screen "Dos" 800x480, template "Main"
   Button "Button_1" at 7,5 size 96x32; TextOff 'Мешалки'; Authorization "Admin"
      on Release: ActivateScreen("Mix", 0); SetTag("settings", 1)
      Appearance <- "settings"
   Button "Button_2" at 7,52 size 96x32; TextOff 'Дозаторы'; Authorization "Admin"
      on Release: ActivateScreen("Dos", 0); SetTag("settings", 2)
      Appearance <- "settings"
   Button "Button_3" at 7,99 size 96x32; TextOff 'Клапана'; Authorization "Admin"
      on Release: ActivateScreen("Valve", 0); SetTag("settings", 3)
      Appearance <- "settings"
   Button "Button_4" at 7,146 size 96x32; TextOff 'AI'; Authorization "Admin"
      on Release: ActivateScreen("AI", 0); SetTag("settings", 4)
      Appearance <- "settings"
   Button "Button_5" at 7,193 size 96x32; TextOff 'DI'; Authorization "Admin"
      on Release: ActivateScreen("DI", 0); SetTag("settings", 5)
      Appearance <- "settings"
   Button "Button_6" at 7,240 size 96x32; TextOff 'DO'; Authorization "Admin"
      on Release: ActivateScreen("DO", 0); SetTag("settings", 6)
      Appearance <- "settings"
   Group "Group" at 127,7 size 416x126; TextList "Hand"; Picture "z2use_3"; PictureList "Motor"; Text 'Мешалка 1'
   Group "Group_1" at 127,146 size 416x126; Text 'Мешалка 1'; PictureList "Motor"; TextList "Hand"; Picture "z2use_3"
   Group "Group_2" at 127,285 size 416x126; Text 'Мешалка 1'; PictureList "Motor"; TextList "Hand"; Picture "z2use_3"
   Rectangle "Rectangle_1" at 127,7 size 416x126
      Appearance <- "Motors_DB_DD_CMD_Sim"
   GraphicIOField "Graphic I/O field_2" at 134,43 size 43x85; PictureList "Motor"
      ProcessValue <- "Motors_DB_DD_Status"
   Button "Button_7" at 213,41 size 90x22; TextOff 'Авто'; TextList "Hand"
      on Click: InvertBit("Motors_DB_DD_CMD_Hand")
      Appearance <- "Motors_DB_DD_CMD_Hand"
      ProcessValue <- "Motors_DB_DD_CMD_Hand"
   Button "Button_8" at 258,63 size 45x22; TextOff 'Выкл'
      on Click: ResetBit("Motors_DB_DD_CMD_Start_M")
   Button "Button_9" at 213,86 size 90x20; TextOff 'Сервис'
      on Click: InvertBit("Motors_DB_DD_CMD_Service")
      Appearance <- "Motors_DB_DD_CMD_Service"
   Button "Button_13" at 213,63 size 45x22; TextOff 'Вкл'
      on Click: SetBit("Motors_DB_DD_CMD_Start_M")
      Appearance <- "Motors_DB_DD_CMD_Start_M"
   TextField "Text field_13" at 133,12 size 171x26; Text 'Сухой дозатор'
   TextField "Text field_15" at 310,12 size 99x18; Text 'Ожидание ОС, с'
   GraphicView "Graphic view_1" at 180,42 size 25x25; Picture "z2use_3"
      Visibility <- "Motors_DB_DD_CMD_Hand"
   GraphicView "Graphic view_8" at 180,74 size 25x25; Picture "force"
      Visibility <- "Motors_DB_DD_CMD_Force"
   GraphicView "Graphic view_11" at 180,103 size 25x25; Picture "service"
      Visibility <- "Motors_DB_DD_CMD_Service"
   TextField "Text field_3" at 436,31 size 20x18; Text 'QF'
   TextField "Text field_10" at 436,56 size 21x18; Text 'KM'
   TextField "Text field_12" at 436,82 size 44x18; Text 'Service'
   TextField "Text field_14" at 436,108 size 41x18; Text 'Termo'
   TextField "Text field_4" at 416,10 size 120x22; Text 'Использовать:'
   Button "Button_21" at 478,32 size 60x20; TextOff 'Text'; Authorization "Operator"; PictureList "ON_OFF"
      on Click: InvertBit("Motors_DB_DD_Use_QF")
      ProcessValue <- "Motors_DB_DD_Use_QF"
   Button "Button_22" at 478,56 size 60x20; TextOff 'Text'; PictureList "ON_OFF"; Authorization "Operator"
      on Click: InvertBit("Motors_DB_DD_Use_KM")
      ProcessValue <- "Motors_DB_DD_Use_KM"
   Button "Button_24" at 478,80 size 60x20; TextOff 'Text'; PictureList "ON_OFF"; Authorization "Operator"
      on Click: InvertBit("Motors_DB_DD_Use_Serivce")
      ProcessValue <- "Motors_DB_DD_Use_Serivce"
   Button "Button_25" at 478,105 size 60x20; TextOff 'Text'; PictureList "ON_OFF"; Authorization "Operator"
      on Click: InvertBit("Motors_DB_DD_Use_Termo")
      ProcessValue <- "Motors_DB_DD_Use_Termo"
   Button "Button_26" at 416,31 size 20x20; TextOff 'Text'; Authorization "Operator"; PictureList "ok"
      ProcessValue <- "Motors_DB_DD_FB_QF"
   Button "Button_27" at 416,55 size 20x20; TextOff 'Text'; PictureList "ok"; Authorization "Operator"
      ProcessValue <- "Motors_DB_DD_FB_KM"
   Button "Button_29" at 416,80 size 20x20; TextOff 'Text'; PictureList "ok"; Authorization "Operator"
      ProcessValue <- "Motors_DB_DD_Use_Serivce"
   Button "Button_30" at 416,105 size 20x20; TextOff 'Text'; PictureList "ok"; Authorization "Operator"
      ProcessValue <- "Motors_DB_DD_FB_Termo"
   TextField "Text field_1" at 323,87 size 79x18; Text 'Наработка, ч'
   TextField "Text field_2" at 309,34 size 37x18; Text 'Старт'
   IOField "I/O field_5" at 348,32 size 30x20; FormatPattern 99
      ProcessValue <- "Motors_DB_DD_Wait_On_SP"
   IOField "I/O field_12" at 348,55 size 30x20; FormatPattern 99
      ProcessValue <- "Motors_DB_DD_Wait_Off_SP"
   TextField "Text field_5" at 309,55 size 32x18; Text 'Стоп'
   IOField "I/O field_13" at 378,32 size 30x20; FormatPattern 99
      ProcessValue <- "Motors_DB_DD_Wait_On_Now"
   IOField "I/O field_14" at 378,55 size 30x20; FormatPattern 99
      ProcessValue <- "Motors_DB_DD_Wait_Off_Now"
   IOField "I/O field_16" at 313,105 size 98x20; FormatPattern 9999999999
      ProcessValue <- "Motors_DB_DD_Res_h"
   Button "Button_11" at 213,106 size 90x20; TextOff 'Force'
      on Click: InvertBit("Motors_DB_DD_CMD_Force")
      Appearance <- "Motors_DB_DD_CMD_Force"
   Rectangle "Rectangle_2" at 127,146 size 416x126
      Appearance <- "Motors_DB_Vibro_CMD_Sim"
   GraphicIOField "Graphic I/O field_1" at 134,182 size 43x85; PictureList "Motor"
      ProcessValue <- "Motors_DB_Vibro_Status"
   Button "Button_10" at 213,180 size 90x22; TextOff 'Авто'; TextList "Hand"
      on Click: InvertBit("Motors_DB_Vibro_CMD_Hand")
      Appearance <- "Motors_DB_Vibro_CMD_Hand"
      ProcessValue <- "Motors_DB_Vibro_CMD_Hand"
   Button "Button_12" at 258,202 size 45x22; TextOff 'Выкл'
      on Click: ResetBit("Motors_DB_Vibro_CMD_Start_M")
   Button "Button_14" at 213,225 size 90x20; TextOff 'Сервис'
      on Click: InvertBit("Motors_DB_Vibro_CMD_Service")
      Appearance <- "Motors_DB_Vibro_CMD_Service"
   Button "Button_15" at 213,202 size 45x22; TextOff 'Вкл'
      on Click: SetBit("Motors_DB_Vibro_CMD_Start_M")
      Appearance <- "Motors_DB_Vibro_CMD_Start_M"
   TextField "Text field_6" at 133,151 size 171x26; Text 'Вибратор'
   TextField "Text field_7" at 310,151 size 99x18; Text 'Ожидание ОС, с'
   GraphicView "Graphic view_2" at 180,181 size 25x25; Picture "z2use_3"
      Visibility <- "Motors_DB_Vibro_CMD_Hand"
   GraphicView "Graphic view_3" at 180,213 size 25x25; Picture "force"
      Visibility <- "Motors_DB_Vibro_CMD_Force"
   GraphicView "Graphic view_4" at 180,242 size 25x25; Picture "service"
      Visibility <- "Motors_DB_Vibro_CMD_Service"
   TextField "Text field_8" at 436,170 size 20x18; Text 'QF'
   TextField "Text field_9" at 436,195 size 21x18; Text 'KM'
   TextField "Text field_11" at 436,221 size 44x18; Text 'Service'
   TextField "Text field_16" at 436,247 size 41x18; Text 'Termo'
   TextField "Text field_17" at 416,149 size 120x22; Text 'Использовать:'
   Button "Button_16" at 478,171 size 60x20; TextOff 'Text'; PictureList "ON_OFF"; Authorization "Operator"
      on Click: InvertBit("Motors_DB_Vibro_Use_QF")
      ProcessValue <- "Motors_DB_Vibro_Use_QF"
   Button "Button_17" at 478,195 size 60x20; TextOff 'Text'; Authorization "Operator"; PictureList "ON_OFF"
      on Click: InvertBit("Motors_DB_Vibro_Use_KM")
      ProcessValue <- "Motors_DB_Vibro_Use_KM"
   Button "Button_18" at 478,219 size 60x20; TextOff 'Text'; Authorization "Operator"; PictureList "ON_OFF"
      on Click: InvertBit("Motors_DB_Vibro_Use_Serivce")
      ProcessValue <- "Motors_DB_Vibro_Use_Serivce"
   Button "Button_19" at 478,244 size 60x20; TextOff 'Text'; Authorization "Operator"; PictureList "ON_OFF"
      on Click: InvertBit("Motors_DB_Vibro_Use_Termo")
      ProcessValue <- "Motors_DB_Vibro_Use_Termo"
   Button "Button_20" at 416,170 size 20x20; TextOff 'Text'; PictureList "ok"; Authorization "Operator"
      ProcessValue <- "Motors_DB_Vibro_FB_QF"
   Button "Button_23" at 416,194 size 20x20; TextOff 'Text'; Authorization "Operator"; PictureList "ok"
      ProcessValue <- "Motors_DB_Vibro_FB_KM"
   Button "Button_28" at 416,219 size 20x20; TextOff 'Text'; Authorization "Operator"; PictureList "ok"
      ProcessValue <- "Motors_DB_Vibro_Use_Serivce"
   Button "Button_31" at 416,244 size 20x20; TextOff 'Text'; Authorization "Operator"; PictureList "ok"
      ProcessValue <- "Motors_DB_Vibro_FB_Termo"
   TextField "Text field_18" at 323,226 size 79x18; Text 'Наработка, ч'
   TextField "Text field_19" at 309,173 size 37x18; Text 'Старт'
   IOField "I/O field_1" at 348,171 size 30x20; FormatPattern 99
      ProcessValue <- "Motors_DB_Vibro_Wait_On_SP"
   IOField "I/O field_2" at 348,194 size 30x20; FormatPattern 99
      ProcessValue <- "Motors_DB_Vibro_Wait_Off_SP"
   TextField "Text field_20" at 309,194 size 32x18; Text 'Стоп'
   IOField "I/O field_3" at 378,171 size 30x20; FormatPattern 99
      ProcessValue <- "Motors_DB_Vibro_Wait_On_Now"
   IOField "I/O field_4" at 378,194 size 30x20; FormatPattern 99
      ProcessValue <- "Motors_DB_Vibro_Wait_Off_Now"
   IOField "I/O field_6" at 313,244 size 98x20; FormatPattern 9999999999
      ProcessValue <- "Motors_DB_Vibro_Res_h"
   Button "Button_32" at 213,245 size 90x20; TextOff 'Force'
      on Click: InvertBit("Motors_DB_Vibro_CMD_Force")
      Appearance <- "Motors_DB_Vibro_CMD_Force"
   Rectangle "Rectangle_3" at 127,285 size 416x126
      Appearance <- "Motors_DB_DL_CMD_Sim"
   GraphicIOField "Graphic I/O field_3" at 134,321 size 43x85; PictureList "Motor"
      ProcessValue <- "Motors_DB_DL_Status"
   Button "Button_33" at 213,319 size 90x22; TextOff 'Авто'; TextList "Hand"
      on Click: InvertBit("Motors_DB_DL_CMD_Hand")
      Appearance <- "Motors_DB_DL_CMD_Hand"
      ProcessValue <- "Motors_DB_DL_CMD_Hand"
   Button "Button_34" at 258,341 size 45x22; TextOff 'Выкл'
      on Click: ResetBit("Motors_DB_DL_CMD_Start_M")
   Button "Button_35" at 213,364 size 90x20; TextOff 'Сервис'
      on Click: InvertBit("Motors_DB_DL_CMD_Service")
      Appearance <- "Motors_DB_DL_CMD_Service"
   Button "Button_36" at 213,341 size 45x22; TextOff 'Вкл'
      on Click: SetBit("Motors_DB_DL_CMD_Start_M")
      Appearance <- "Motors_DB_DL_CMD_Start_M"
   TextField "Text field_21" at 133,290 size 171x26; Text 'Жидкий дозатор'
   TextField "Text field_22" at 310,290 size 99x18; Text 'Ожидание ОС, с'
   GraphicView "Graphic view_5" at 180,320 size 25x25; Picture "z2use_3"
      Visibility <- "Motors_DB_DL_CMD_Hand"
   GraphicView "Graphic view_6" at 180,352 size 25x25; Picture "force"
      Visibility <- "Motors_DB_DL_CMD_Force"
   GraphicView "Graphic view_7" at 180,381 size 25x25; Picture "service"
      Visibility <- "Motors_DB_DL_CMD_Service"
   TextField "Text field_23" at 436,309 size 20x18; Text 'QF'
   TextField "Text field_24" at 436,334 size 21x18; Text 'KM'
   TextField "Text field_25" at 436,360 size 44x18; Text 'Service'
   TextField "Text field_26" at 436,386 size 41x18; Text 'Termo'
   TextField "Text field_27" at 416,288 size 120x22; Text 'Использовать:'
   Button "Button_37" at 478,310 size 60x20; TextOff 'Text'; PictureList "ON_OFF"; Authorization "Operator"
      on Click: InvertBit("Motors_DB_DL_Use_QF")
      ProcessValue <- "Motors_DB_DL_Use_QF"
   Button "Button_38" at 478,334 size 60x20; TextOff 'Text'; Authorization "Operator"; PictureList "ON_OFF"
      on Click: InvertBit("Motors_DB_DL_Use_KM")
      ProcessValue <- "Motors_DB_DL_Use_KM"
   Button "Button_39" at 478,358 size 60x20; TextOff 'Text'; Authorization "Operator"; PictureList "ON_OFF"
      on Click: InvertBit("Motors_DB_DL_Use_Serivce")
      ProcessValue <- "Motors_DB_DL_Use_Serivce"
   Button "Button_40" at 478,383 size 60x20; TextOff 'Text'; Authorization "Operator"; PictureList "ON_OFF"
      on Click: InvertBit("Motors_DB_DL_Use_Termo")
      ProcessValue <- "Motors_DB_DL_Use_Termo"
   Button "Button_41" at 416,309 size 20x20; TextOff 'Text'; PictureList "ok"; Authorization "Operator"
      ProcessValue <- "Motors_DB_DL_FB_QF"
   Button "Button_42" at 416,333 size 20x20; TextOff 'Text'; Authorization "Operator"; PictureList "ok"
      ProcessValue <- "Motors_DB_DL_FB_KM"
   Button "Button_43" at 416,358 size 20x20; TextOff 'Text'; Authorization "Operator"; PictureList "ok"
      ProcessValue <- "Motors_DB_DL_Use_Serivce"
   Button "Button_44" at 416,383 size 20x20; TextOff 'Text'; Authorization "Operator"; PictureList "ok"
      ProcessValue <- "Motors_DB_DL_FB_Termo"
   TextField "Text field_28" at 323,365 size 79x18; Text 'Наработка, ч'
   TextField "Text field_29" at 309,312 size 37x18; Text 'Старт'
   IOField "I/O field_7" at 348,310 size 30x20; FormatPattern 99
      ProcessValue <- "Motors_DB_DL_Wait_On_SP"
   IOField "I/O field_8" at 348,333 size 30x20; FormatPattern 99
      ProcessValue <- "Motors_DB_DL_Wait_Off_SP"
   TextField "Text field_30" at 309,333 size 32x18; Text 'Стоп'
   IOField "I/O field_9" at 378,310 size 30x20; FormatPattern 99
      ProcessValue <- "Motors_DB_DL_Wait_On_Now"
   IOField "I/O field_10" at 378,333 size 30x20; FormatPattern 99
      ProcessValue <- "Motors_DB_DL_Wait_Off_Now"
   IOField "I/O field_11" at 313,383 size 98x20; FormatPattern 9999999999
      ProcessValue <- "Motors_DB_DL_Res_h"
   Button "Button_45" at 213,384 size 90x20; TextOff 'Force'
      on Click: InvertBit("Motors_DB_DL_CMD_Force")
      Appearance <- "Motors_DB_DL_CMD_Force"

screen "Valve" 800x480, template "Main"
   Button "Button_1" at 7,5 size 96x32; TextOff 'Мешалки'; Authorization "Admin"
      on Release: ActivateScreen("Mix", 0); SetTag("settings", 1)
      Appearance <- "settings"
   Button "Button_2" at 7,52 size 96x32; TextOff 'Дозаторы'; Authorization "Admin"
      on Release: ActivateScreen("Dos", 0); SetTag("settings", 2)
      Appearance <- "settings"
   Button "Button_3" at 7,99 size 96x32; TextOff 'Клапана'; Authorization "Admin"
      on Release: ActivateScreen("Valve", 0); SetTag("settings", 3)
      Appearance <- "settings"
   Button "Button_4" at 7,146 size 96x32; TextOff 'AI'; Authorization "Admin"
      on Release: ActivateScreen("AI", 0); SetTag("settings", 4)
      Appearance <- "settings"
   Button "Button_5" at 7,193 size 96x32; TextOff 'DI'; Authorization "Admin"
      on Release: ActivateScreen("DI", 0); SetTag("settings", 5)
      Appearance <- "settings"
   Button "Button_6" at 7,240 size 96x32; TextOff 'DO'; Authorization "Admin"
      on Release: ActivateScreen("DO", 0); SetTag("settings", 6)
      Appearance <- "settings"
   Group "Group" at 127,7 size 264x51; TextList "Hand"
   Rectangle "Rectangle_2" at 127,7 size 264x51
      Appearance <- "Micro_DB_KC1_Alarm"
   TextField "Text field_5" at 130,10 size 97x22; Text 'Клапан КС1'
   Button "Button_13" at 246,11 size 59x44; TextOff 'Авто'; TextList "Hand"
      on Click: InvertBit("Micro_DB_KC1_Hand")
      Appearance <- "Micro_DB_KC1_Hand"
      ProcessValue <- "Micro_DB_KC1_Hand"
   Button "Button_14" at 188,33 size 49x22; TextOff 'Выкл'
      on Click: ResetBit("Micro_DB_KC1_Start_M")
   Button "Button_15" at 132,33 size 47x22; TextOff 'Вкл'
      on Click: SetBit("Micro_DB_KC1_Start_M")
      Appearance <- "Micro_DB_KC1_Start_M"
   TextField "Text field_1" at 306,8 size 28x23; Text 'ОС'
   Button "Button_7" at 336,11 size 50x20; TextOff 'Text'; Authorization "Operator"; PictureList "ON_OFF"
      on Click: InvertBit("Micro_DB_KC1_No_FB")
      ProcessValue <- "Micro_DB_KC1_No_FB"
   IOField "I/O field_5" at 308,31 size 30x22; FormatPattern 99
      ProcessValue <- "Micro_DB_KC1_Wait_On_SP"
   IOField "I/O field_8" at 355,31 size 30x22; FormatPattern 99
      ProcessValue <- "Micro_DB_KC1_Wait_Off_SP"

screen "AI" 800x480, template "Main"
   Button "Button_1" at 7,5 size 96x32; TextOff 'Мешалки'; Authorization "Admin"
      on Release: ActivateScreen("Mix", 0); SetTag("settings", 1)
      Appearance <- "settings"
   Button "Button_2" at 7,52 size 96x32; TextOff 'Дозаторы'; Authorization "Admin"
      on Release: ActivateScreen("Dos", 0); SetTag("settings", 2)
      Appearance <- "settings"
   Button "Button_3" at 7,99 size 96x32; TextOff 'Клапана'; Authorization "Admin"
      on Release: ActivateScreen("Valve", 0); SetTag("settings", 3)
      Appearance <- "settings"
   Button "Button_4" at 7,146 size 96x32; TextOff 'AI'; Authorization "Admin"
      on Release: ActivateScreen("AI", 0); SetTag("settings", 4)
      Appearance <- "settings"
   Button "Button_5" at 7,193 size 96x32; TextOff 'DI'; Authorization "Admin"
      on Release: ActivateScreen("DI", 0); SetTag("settings", 5)
      Appearance <- "settings"
   Button "Button_6" at 7,240 size 96x32; TextOff 'DO'; Authorization "Admin"
      on Release: ActivateScreen("DO", 0); SetTag("settings", 6)
      Appearance <- "settings"
   TextField "Text field_2" at 210,15 size 67x22; Text 'Датчик:'
   TextField "Text field_4" at 282,15 size 99x22; Text 'Расходомер'
   TextField "Text field_7" at 390,18 size 43x22; Text 'вход'
   TextField "Text field_8" at 390,43 size 56x22; Text 'выход'
   IOField "I/O field_1" at 456,19 size 92x26; FormatPattern s999999999.999
      ProcessValue <- "AIx_DB_FlowMeter_Converter_Min_In"
   IOField "I/O field_2" at 456,41 size 92x26; FormatPattern s999999999.999
      ProcessValue <- "AIx_DB_FlowMeter_Converter_Min_Out"
   IOField "I/O field_3" at 555,18 size 92x26; FormatPattern s999999999.999
      ProcessValue <- "AIx_DB_FlowMeter_Converter_Max_In"
   IOField "I/O field_4" at 555,40 size 92x26; FormatPattern s999999999.999
      ProcessValue <- "AIx_DB_FlowMeter_Converter_Max_Out"
   TextField "Text field_9" at 389,68 size 101x22; Text 'Фильтрация'
   TextField "Text field_10" at 390,96 size 36x22; Text 'RTD'
   Button "Button_7" at 489,71 size 20x20; TextOff 'Text'; PictureList "ok"
      ProcessValue <- "AIx_DB_FlowMeter_Use_Filter"
      on Click: InvertBit("AIx_DB_FlowMeter_Use_Filter")
   Button "Button_8" at 489,96 size 20x20; TextOff 'Text'; PictureList "ok"
      on Click: InvertBit("AIx_DB_FlowMeter_Use_RTD")
      ProcessValue <- "AIx_DB_FlowMeter_Use_RTD"
   IOField "I/O field_5" at 516,68 size 65x25; FormatPattern 999
      ProcessValue <- "AIx_DB_FlowMeter_Filter_SP"
   IOField "I/O field_6" at 516,93 size 65x25; FormatPattern 999
      ProcessValue <- "AIx_DB_FlowMeter_RTD_c"
   TextField "Text field_11" at 210,36 size 79x22; Text 'Поправка'
   IOField "I/O field_7" at 293,36 size 78x23; FormatPattern s999.9
      ProcessValue <- "AIx_DB_FlowMeter_Calibration"
   Button "Button_9" at 396,176 size 248x28; TextOff 'Use'
      Appearance <- "AIx_DB_FlowMeter_CMD_Start_A"
      on Click: InvertBit("AIx_DB_FlowMeter_CMD_Start_A")
   Button "Button_10" at 213,66 size 68x28; TextOff 'Hand'
      on Click: InvertBit("AIx_DB_FlowMeter_CMD_Hand")
      Appearance <- "AIx_DB_FlowMeter_CMD_Hand"
   IOField "I/O field_8" at 293,66 size 78x28; FormatPattern s9999.9
      ProcessValue <- "AIx_DB_FlowMeter_Result"
   TextField "Text field_12" at 436,123 size 27x22; Text 'NC'
   TextField "Text field_13" at 437,143 size 25x22; Text 'SC'
   TextField "Text field_14" at 210,125 size 27x22; Text 'HH'
   TextField "Text field_15" at 216,145 size 16x22; Text 'H'
   TextField "Text field_16" at 217,165 size 14x22; Text 'L'
   TextField "Text field_17" at 212,186 size 23x22; Text 'LL'
   IOField "I/O field_11" at 472,123 size 58x21; FormatPattern s99999
      ProcessValue <- "AIx_DB_FlowMeter_SP_NC"
   IOField "I/O field_12" at 472,143 size 58x21; FormatPattern s99999
      ProcessValue <- "AIx_DB_FlowMeter_SP_SC"
   IOField "I/O field_13" at 246,125 size 58x21; FormatPattern 99999
      ProcessValue <- "AIx_DB_FlowMeter_SP_HH"
   IOField "I/O field_14" at 246,145 size 58x21; FormatPattern 99999
      ProcessValue <- "AIx_DB_FlowMeter_SP_H"
   IOField "I/O field_15" at 246,165 size 58x21; FormatPattern s99999
      ProcessValue <- "AIx_DB_FlowMeter_SP_L"
   IOField "I/O field_16" at 246,185 size 58x21; FormatPattern s99999
      ProcessValue <- "AIx_DB_FlowMeter_SP_LL"
   IOField "I/O field_17" at 546,123 size 58x21; FormatPattern 999
      ProcessValue <- "AIx_DB_FlowMeter_Timers_NC_SP"
   IOField "I/O field_18" at 546,143 size 58x21; FormatPattern 999
      ProcessValue <- "AIx_DB_FlowMeter_Timers_SC_SP"
   IOField "I/O field_19" at 320,125 size 58x21; FormatPattern 999
      ProcessValue <- "AIx_DB_FlowMeter_Timers_HH_SP"
   IOField "I/O field_20" at 320,145 size 58x21; FormatPattern 999
      ProcessValue <- "AIx_DB_FlowMeter_Timers_H_SP"
   IOField "I/O field_21" at 320,165 size 58x21; FormatPattern 999
      ProcessValue <- "AIx_DB_FlowMeter_Timers_L_SP"
   IOField "I/O field_22" at 320,185 size 58x21; FormatPattern 999
      ProcessValue <- "AIx_DB_FlowMeter_Timers_LL_SP"
   IOField "I/O field_23" at 582,93 size 65x25; FormatPattern s99999
      ProcessValue <- "AIx_DB_FlowMeter_Signal"
   TextField "Text field_18" at 210,97 size 68x22; Text 'Уставка'
   TextField "Text field_19" at 299,97 size 79x22; Text 'Время (с)'
   TextField "Text field_1" at 214,248 size 67x22; Text 'Датчик:'
   TextField "Text field_3" at 286,248 size 69x22; Text 'Уровень'
   TextField "Text field_5" at 394,251 size 43x22; Text 'вход'
   TextField "Text field_6" at 394,276 size 56x22; Text 'выход'
   IOField "I/O field_9" at 460,252 size 92x26; FormatPattern s999999999.999
      ProcessValue <- "AIx_DB_Level_Converter_Min_In"
   IOField "I/O field_10" at 460,274 size 92x26; FormatPattern s999999999.999
      ProcessValue <- "AIx_DB_Level_Converter_Min_Out"
   IOField "I/O field_24" at 559,251 size 92x26; FormatPattern s999999999.999
      ProcessValue <- "AIx_DB_Level_Converter_Max_In"
   IOField "I/O field_25" at 559,273 size 92x26; FormatPattern s999999999.999
      ProcessValue <- "AIx_DB_Level_Converter_Max_Out"
   TextField "Text field_20" at 393,301 size 101x22; Text 'Фильтрация'
   TextField "Text field_21" at 394,329 size 36x22; Text 'RTD'
   Button "Button_11" at 493,304 size 20x20; TextOff 'Text'; PictureList "ok"
      on Click: InvertBit("AIx_DB_Level_Use_Filter")
      ProcessValue <- "AIx_DB_Level_Use_Filter"
   Button "Button_12" at 493,329 size 20x20; TextOff 'Text'; PictureList "ok"
      on Click: InvertBit("AIx_DB_Level_Use_RTD")
      ProcessValue <- "AIx_DB_Level_Use_RTD"
   IOField "I/O field_26" at 520,301 size 65x25; FormatPattern 999
      ProcessValue <- "AIx_DB_Level_Filter_SP"
   IOField "I/O field_27" at 520,326 size 65x25; FormatPattern 999
      ProcessValue <- "AIx_DB_Level_RTD_c"
   TextField "Text field_22" at 214,269 size 79x22; Text 'Поправка'
   IOField "I/O field_28" at 297,269 size 78x23; FormatPattern s999.9
      ProcessValue <- "AIx_DB_Level_Calibration"
   Button "Button_13" at 400,409 size 248x28; TextOff 'Use'
      on Click: InvertBit("AIx_DB_Level_CMD_Start_A")
      Appearance <- "AIx_DB_Level_CMD_Start_A"
   Button "Button_14" at 217,299 size 68x28; TextOff 'Hand'
      on Click: InvertBit("AIx_DB_Level_CMD_Hand")
      Appearance <- "AIx_DB_Level_CMD_Hand"
   IOField "I/O field_29" at 297,299 size 78x28; FormatPattern s9999.9
      ProcessValue <- "AIx_DB_Level_Result"
   TextField "Text field_23" at 440,356 size 27x22; Text 'NC'
   TextField "Text field_24" at 441,376 size 25x22; Text 'SC'
   TextField "Text field_25" at 214,358 size 27x22; Text 'HH'
   TextField "Text field_26" at 220,378 size 16x22; Text 'H'
   TextField "Text field_27" at 221,398 size 14x22; Text 'L'
   TextField "Text field_28" at 216,419 size 23x22; Text 'LL'
   IOField "I/O field_30" at 476,356 size 58x21; FormatPattern s99999
      ProcessValue <- "AIx_DB_Level_SP_NC"
   IOField "I/O field_31" at 476,376 size 58x21; FormatPattern s99999
      ProcessValue <- "AIx_DB_Level_SP_SC"
   IOField "I/O field_32" at 250,358 size 58x21; FormatPattern 99999
      ProcessValue <- "AIx_DB_Level_SP_HH"
   IOField "I/O field_33" at 250,378 size 58x21; FormatPattern 99999
      ProcessValue <- "AIx_DB_Level_SP_H"
   IOField "I/O field_34" at 250,398 size 58x21; FormatPattern s99999
      ProcessValue <- "AIx_DB_Level_SP_L"
   IOField "I/O field_35" at 250,418 size 58x21; FormatPattern s99999
      ProcessValue <- "AIx_DB_Level_SP_LL"
   IOField "I/O field_36" at 550,356 size 58x21; FormatPattern 999
      ProcessValue <- "AIx_DB_Level_Timers_NC_SP"
   IOField "I/O field_37" at 550,376 size 58x21; FormatPattern 999
      ProcessValue <- "AIx_DB_Level_Timers_SC_SP"
   IOField "I/O field_38" at 324,358 size 58x21; FormatPattern 999
      ProcessValue <- "AIx_DB_Level_Timers_HH_SP"
   IOField "I/O field_39" at 324,378 size 58x21; FormatPattern 999
      ProcessValue <- "AIx_DB_Level_Timers_H_SP"
   IOField "I/O field_40" at 324,398 size 58x21; FormatPattern 999
      ProcessValue <- "AIx_DB_Level_Timers_L_SP"
   IOField "I/O field_41" at 324,418 size 58x21; FormatPattern 999
      ProcessValue <- "AIx_DB_Level_Timers_LL_SP"
   IOField "I/O field_42" at 586,326 size 65x25; FormatPattern s99999
      ProcessValue <- "AIx_DB_Level_Signal"
   TextField "Text field_29" at 214,330 size 68x22; Text 'Уставка'
   TextField "Text field_30" at 303,330 size 79x22; Text 'Время (с)'

screen "DI" 800x480, template "Main"
   Button "Button_1" at 7,5 size 96x32; TextOff 'Мешалки'; Authorization "Admin"
      on Release: ActivateScreen("Mix", 0); SetTag("settings", 1)
      Appearance <- "settings"
   Button "Button_2" at 7,52 size 96x32; TextOff 'Дозаторы'; Authorization "Admin"
      on Release: ActivateScreen("Dos", 0); SetTag("settings", 2)
      Appearance <- "settings"
   Button "Button_3" at 7,99 size 96x32; TextOff 'Клапана'; Authorization "Admin"
      on Release: ActivateScreen("Valve", 0); SetTag("settings", 3)
      Appearance <- "settings"
   Button "Button_4" at 7,146 size 96x32; TextOff 'AI'; Authorization "Admin"
      on Release: ActivateScreen("AI", 0); SetTag("settings", 4)
      Appearance <- "settings"
   Button "Button_5" at 7,193 size 96x32; TextOff 'DI'; Authorization "Admin"
      on Release: ActivateScreen("DI", 0); SetTag("settings", 5)
      Appearance <- "settings"
   Button "Button_6" at 7,240 size 96x32; TextOff 'DO'; Authorization "Admin"
      on Release: ActivateScreen("DO", 0); SetTag("settings", 6)
      Appearance <- "settings"
   Group "Group" at 127,7 size 283x51; TextList "Hand"
   Group "Group_1" at 127,66 size 283x51; TextList "Hand"
   Group "Group_2" at 127,125 size 283x51; TextList "Hand"
   Group "Group_3" at 127,184 size 283x51; TextList "Hand"
   Group "Group_4" at 127,244 size 283x51; TextList "Hand"
   Group "Group_5" at 127,303 size 283x51; TextList "Hand"
   Group "Group_6" at 127,362 size 283x51; TextList "Hand"
   Group "Group_7" at 127,422 size 283x51; TextList "Hand"
   Group "Group_8" at 433,7 size 283x51; TextList "Hand"
   Group "Group_9" at 433,66 size 283x51; TextList "Hand"
   Group "Group_10" at 433,125 size 283x51; TextList "Hand"
   Group "Group_11" at 433,184 size 283x51; TextList "Hand"
   Group "Group_12" at 433,244 size 283x51; TextList "Hand"
   Group "Group_13" at 433,303 size 283x51; TextList "Hand"
   TextField "Text field_1" at 131,10 size 45x22; Text 'I 0.0'
   TextField "Text field_2" at 176,10 size 120x22; Text 'M1 Готовность'
   Circle "Circle_1" at 131,33 size 22x22
      Appearance <- "DIx_DB_M1_FB_Ready_Input"
   Circle "Circle_2" at 154,33 size 22x22
      Appearance <- "DIx_DB_M1_FB_Ready_Signal"
   Button "Button_7" at 298,11 size 59x44; TextOff 'Авто'; TextList "Hand"
      on Click: InvertBit("DIx_DB_M1_FB_Ready_Hand")
      Appearance <- "DIx_DB_M1_FB_Ready_Hand"
      ProcessValue <- "DIx_DB_M1_FB_Ready_Hand"
   Button "Button_8" at 240,33 size 49x22; TextOff 'Выкл'
      on Click: ResetBit("DIx_DB_M1_FB_Ready_Start_M")
   Button "Button_12" at 184,33 size 47x22; TextOff 'Вкл'
      Appearance <- "DIx_DB_M1_FB_Ready_Start_M"
      on Click: SetBit("DIx_DB_M1_FB_Ready_Start_M")
   IOField "I/O field_6" at 360,33 size 23x22; FormatPattern 99
      ProcessValue <- "DIx_DB_M1_FB_Ready_Filter_On_SP"
   IOField "I/O field_7" at 383,33 size 23x22; FormatPattern 99
      ProcessValue <- "DIx_DB_M1_FB_Ready_Filter_Off_SP"
   Button "Button_9" at 360,10 size 46x20; TextOff 'Inv'
      Appearance <- "DIx_DB_M1_FB_Ready_Inverse"
      on Click: InvertBit("DIx_DB_M1_FB_Ready_Inverse")
   TextField "Text field_3" at 131,69 size 45x22; Text 'I 0.1'
   TextField "Text field_4" at 176,69 size 87x22; Text 'M1 Работа'
   Circle "Circle_3" at 131,92 size 22x22
      Appearance <- "DIx_DB_M1_FB_Run_Input"
   Circle "Circle_4" at 154,92 size 22x22
      Appearance <- "DIx_DB_M1_FB_Run_Signal"
   Button "Button_10" at 298,70 size 59x44; TextOff 'Авто'; TextList "Hand"
      on Click: InvertBit("DIx_DB_M1_FB_Run_Hand")
      Appearance <- "DIx_DB_M1_FB_Run_Hand"
      ProcessValue <- "DIx_DB_M1_FB_Run_Hand"
   Button "Button_11" at 240,92 size 49x22; TextOff 'Выкл'
      on Click: ResetBit("DIx_DB_M1_FB_Run_Start_M")
   Button "Button_13" at 184,92 size 47x22; TextOff 'Вкл'
      on Click: SetBit("DIx_DB_M1_FB_Run_Start_M")
      Appearance <- "DIx_DB_M1_FB_Run_Start_M"
   IOField "I/O field_1" at 360,92 size 23x22; FormatPattern 99
      ProcessValue <- "DIx_DB_M1_FB_Run_Filter_On_SP"
   IOField "I/O field_2" at 383,92 size 23x22; FormatPattern 99
      ProcessValue <- "DIx_DB_M1_FB_Run_Filter_Off_SP"
   Button "Button_14" at 360,69 size 46x20; TextOff 'Inv'
      on Click: InvertBit("DIx_DB_M1_FB_Run_Inverse")
      Appearance <- "DIx_DB_M1_FB_Run_Inverse"
   TextField "Text field_5" at 131,128 size 45x22; Text 'I 0.2'
   TextField "Text field_6" at 176,128 size 120x22; Text 'M2 Готовность'
   Circle "Circle_5" at 131,151 size 22x22
      Appearance <- "DIx_DB_M2_FB_Ready_Input"
   Circle "Circle_6" at 154,151 size 22x22
      Appearance <- "DIx_DB_M2_FB_Ready_Signal"
   Button "Button_15" at 298,129 size 59x44; TextOff 'Авто'; TextList "Hand"
      on Click: InvertBit("DIx_DB_M2_FB_Ready_Hand")
      Appearance <- "DIx_DB_M2_FB_Ready_Hand"
      ProcessValue <- "DIx_DB_M2_FB_Ready_Hand"
   Button "Button_16" at 240,151 size 49x22; TextOff 'Выкл'
      on Click: ResetBit("DIx_DB_M2_FB_Ready_Start_M")
   Button "Button_17" at 184,151 size 47x22; TextOff 'Вкл'
      on Click: SetBit("DIx_DB_M2_FB_Ready_Start_M")
      Appearance <- "DIx_DB_M2_FB_Ready_Start_M"
   IOField "I/O field_3" at 360,151 size 23x22; FormatPattern 99
      ProcessValue <- "DIx_DB_M2_FB_Ready_Filter_On_SP"
   IOField "I/O field_4" at 383,151 size 23x22; FormatPattern 99
      ProcessValue <- "DIx_DB_M2_FB_Ready_Filter_Off_SP"
   Button "Button_18" at 360,128 size 46x20; TextOff 'Inv'
      on Click: InvertBit("DIx_DB_M2_FB_Ready_Inverse")
      Appearance <- "DIx_DB_M2_FB_Ready_Inverse"
   TextField "Text field_7" at 131,187 size 45x22; Text 'I 0.3'
   TextField "Text field_8" at 176,187 size 87x22; Text 'M2 Работа'
   Circle "Circle_7" at 131,210 size 22x22
      Appearance <- "DIx_DB_M2_FB_Run_Input"
   Circle "Circle_8" at 154,210 size 22x22
      Appearance <- "DIx_DB_M2_FB_Run_Signal"
   Button "Button_19" at 298,188 size 59x44; TextOff 'Авто'; TextList "Hand"
      on Click: InvertBit("DIx_DB_M2_FB_Run_Hand")
      Appearance <- "DIx_DB_M2_FB_Run_Hand"
      ProcessValue <- "DIx_DB_M2_FB_Run_Hand"
   Button "Button_20" at 240,210 size 49x22; TextOff 'Выкл'
      on Click: ResetBit("DIx_DB_M2_FB_Run_Start_M")
   Button "Button_21" at 184,210 size 47x22; TextOff 'Вкл'
      on Click: SetBit("DIx_DB_M2_FB_Run_Start_M")
      Appearance <- "DIx_DB_M2_FB_Run_Start_M"
   IOField "I/O field_5" at 360,210 size 23x22; FormatPattern 99
      ProcessValue <- "DIx_DB_M2_FB_Run_Filter_On_SP"
   IOField "I/O field_8" at 383,210 size 23x22; FormatPattern 99
      ProcessValue <- "DIx_DB_M2_FB_Run_Filter_Off_SP"
   Button "Button_22" at 360,187 size 46x20; TextOff 'Inv'
      on Click: InvertBit("DIx_DB_M2_FB_Run_Inverse")
      Appearance <- "DIx_DB_M2_FB_Run_Inverse"
   TextField "Text field_9" at 131,247 size 45x22; Text 'I 0.4'
   TextField "Text field_10" at 176,247 size 120x22; Text 'M3 Готовность'
   Circle "Circle_9" at 131,270 size 22x22
      Appearance <- "DIx_DB_M3_FB_Ready_Input"
   Circle "Circle_10" at 154,270 size 22x22
      Appearance <- "DIx_DB_M3_FB_Ready_Signal"
   Button "Button_23" at 298,248 size 59x44; TextOff 'Авто'; TextList "Hand"
      on Click: InvertBit("DIx_DB_M3_FB_Ready_Hand")
      Appearance <- "DIx_DB_M3_FB_Ready_Hand"
      ProcessValue <- "DIx_DB_M3_FB_Ready_Hand"
   Button "Button_24" at 240,270 size 49x22; TextOff 'Выкл'
      on Click: ResetBit("DIx_DB_M3_FB_Ready_Start_M")
   Button "Button_25" at 184,270 size 47x22; TextOff 'Вкл'
      on Click: SetBit("DIx_DB_M3_FB_Ready_Start_M")
      Appearance <- "DIx_DB_M3_FB_Ready_Start_M"
   IOField "I/O field_9" at 360,270 size 23x22; FormatPattern 99
      ProcessValue <- "DIx_DB_M3_FB_Ready_Filter_On_SP"
   IOField "I/O field_10" at 383,270 size 23x22; FormatPattern 99
      ProcessValue <- "DIx_DB_M3_FB_Ready_Filter_Off_SP"
   Button "Button_26" at 360,247 size 46x20; TextOff 'Inv'
      on Click: InvertBit("DIx_DB_M3_FB_Ready_Inverse")
      Appearance <- "DIx_DB_M3_FB_Ready_Inverse"
   TextField "Text field_11" at 131,306 size 45x22; Text 'I 0.5'
   TextField "Text field_12" at 176,306 size 87x22; Text 'M3 Работа'
   Circle "Circle_11" at 131,329 size 22x22
      Appearance <- "DIx_DB_M3_FB_Run_Input"
   Circle "Circle_12" at 154,329 size 22x22
      Appearance <- "DIx_DB_M3_FB_Run_Signal"
   Button "Button_27" at 298,307 size 59x44; TextOff 'Авто'; TextList "Hand"
      on Click: InvertBit("DIx_DB_M3_FB_Run_Hand")
      Appearance <- "DIx_DB_M3_FB_Run_Hand"
      ProcessValue <- "DIx_DB_M3_FB_Run_Hand"
   Button "Button_28" at 240,329 size 49x22; TextOff 'Выкл'
      on Click: ResetBit("DIx_DB_M3_FB_Run_Start_M")
   Button "Button_29" at 184,329 size 47x22; TextOff 'Вкл'
      on Click: SetBit("DIx_DB_M3_FB_Run_Start_M")
      Appearance <- "DIx_DB_M3_FB_Run_Start_M"
   IOField "I/O field_11" at 360,329 size 23x22; FormatPattern 99
      ProcessValue <- "DIx_DB_M3_FB_Run_Filter_On_SP"
   IOField "I/O field_12" at 383,329 size 23x22; FormatPattern 99
      ProcessValue <- "DIx_DB_M3_FB_Run_Filter_Off_SP"
   Button "Button_30" at 360,306 size 46x20; TextOff 'Inv'
      on Click: InvertBit("DIx_DB_M3_FB_Run_Inverse")
      Appearance <- "DIx_DB_M3_FB_Run_Inverse"
   TextField "Text field_13" at 131,365 size 45x22; Text 'I 0.6'
   TextField "Text field_14" at 176,365 size 120x22; Text 'Сух.доз.Готов.'
   Circle "Circle_13" at 131,388 size 22x22
      Appearance <- "DIx_DB_DD_FB_Ready_Input"
   Circle "Circle_14" at 154,388 size 22x22
      Appearance <- "DIx_DB_DD_FB_Ready_Signal"
   Button "Button_31" at 298,366 size 59x44; TextOff 'Авто'; TextList "Hand"
      on Click: InvertBit("DIx_DB_DD_FB_Ready_Hand")
      Appearance <- "DIx_DB_DD_FB_Ready_Hand"
      ProcessValue <- "DIx_DB_DD_FB_Ready_Hand"
   Button "Button_32" at 240,388 size 49x22; TextOff 'Выкл'
      on Click: ResetBit("DIx_DB_DD_FB_Ready_Start_M")
   Button "Button_33" at 184,388 size 47x22; TextOff 'Вкл'
      on Click: SetBit("DIx_DB_DD_FB_Ready_Start_M")
      Appearance <- "DIx_DB_DD_FB_Ready_Start_M"
   IOField "I/O field_13" at 360,388 size 23x22; FormatPattern 99
      ProcessValue <- "DIx_DB_DD_FB_Ready_Filter_On_SP"
   IOField "I/O field_14" at 383,388 size 23x22; FormatPattern 99
      ProcessValue <- "DIx_DB_DD_FB_Ready_Filter_Off_SP"
   Button "Button_34" at 360,365 size 46x20; TextOff 'Inv'
      on Click: InvertBit("DIx_DB_DD_FB_Ready_Inverse")
      Appearance <- "DIx_DB_DD_FB_Ready_Inverse"
   TextField "Text field_15" at 131,425 size 45x22; Text 'I 0.7'
   TextField "Text field_16" at 176,425 size 98x22; Text 'Доз. Работа'
   Circle "Circle_15" at 131,448 size 22x22
      Appearance <- "DIx_DB_Dos_FB_Run_Input"
   Circle "Circle_16" at 154,448 size 22x22
      Appearance <- "DIx_DB_Dos_FB_Run_Signal"
   Button "Button_35" at 298,426 size 59x44; TextOff 'Авто'; TextList "Hand"
      on Click: InvertBit("DIx_DB_Dos_FB_Run_Hand")
      ProcessValue <- "DIx_DB_Dos_FB_Run_Hand"
      Appearance <- "DIx_DB_Dos_FB_Run_Hand"
   Button "Button_36" at 240,448 size 49x22; TextOff 'Выкл'
      on Click: ResetBit("DIx_DB_Dos_FB_Run_Start_M")
   Button "Button_37" at 184,448 size 47x22; TextOff 'Вкл'
      on Click: SetBit("DIx_DB_Dos_FB_Run_Start_M")
      Appearance <- "DIx_DB_Dos_FB_Run_Start_M"
   IOField "I/O field_15" at 360,448 size 23x22; FormatPattern 99
      ProcessValue <- "DIx_DB_Dos_FB_Run_Filter_On_SP"
   IOField "I/O field_16" at 383,448 size 23x22; FormatPattern 99
      ProcessValue <- "DIx_DB_Dos_FB_Run_Filter_Off_SP"
   Button "Button_38" at 360,425 size 46x20; TextOff 'Inv'
      on Click: InvertBit("DIx_DB_Dos_FB_Run_Inverse")
      Appearance <- "DIx_DB_Dos_FB_Run_Inverse"
   TextField "Text field_17" at 437,10 size 45x22; Text 'I 1.0'
   TextField "Text field_18" at 482,10 size 95x22; Text 'Сух.доз.Ур.'
   Circle "Circle_17" at 437,33 size 22x22
      Appearance <- "DIx_DB_DD_LLS_Input"
   Circle "Circle_18" at 460,33 size 22x22
      Appearance <- "DIx_DB_DD_LLS_Signal"
   Button "Button_39" at 604,11 size 59x44; TextOff 'Авто'; TextList "Hand"
      on Click: InvertBit("DIx_DB_DD_LLS_Hand")
      Appearance <- "DIx_DB_DD_LLS_Hand"
      ProcessValue <- "DIx_DB_DD_LLS_Hand"
   Button "Button_40" at 546,33 size 49x22; TextOff 'Выкл'
      on Click: ResetBit("DIx_DB_DD_LLS_Start_M")
   Button "Button_41" at 490,33 size 47x22; TextOff 'Вкл'
      on Click: SetBit("DIx_DB_DD_LLS_Start_M")
      Appearance <- "DIx_DB_DD_LLS_Start_M"
   IOField "I/O field_17" at 666,33 size 23x22; FormatPattern 99
      ProcessValue <- "DIx_DB_DD_LLS_Filter_On_SP"
   IOField "I/O field_18" at 689,33 size 23x22; FormatPattern 99
      ProcessValue <- "DIx_DB_DD_LLS_Filter_Off_SP"
   Button "Button_42" at 666,10 size 46x20; TextOff 'Inv'
      on Click: InvertBit("DIx_DB_DD_LLS_Inverse")
      Appearance <- "DIx_DB_DD_LLS_Inverse"
   TextField "Text field_19" at 437,69 size 45x22; Text 'I 1.1'
   TextField "Text field_20" at 482,69 size 104x22; Text 'Вибро Готов.'
   Circle "Circle_19" at 437,92 size 22x22
      Appearance <- "DIx_DB_Vibro_FB_Ready_Input"
   Circle "Circle_20" at 460,92 size 22x22
      Appearance <- "DIx_DB_Vibro_FB_Ready_Signal"
   Button "Button_43" at 604,70 size 59x44; TextOff 'Авто'; TextList "Hand"
      on Click: InvertBit("DIx_DB_Vibro_FB_Ready_Hand")
      Appearance <- "DIx_DB_Vibro_FB_Ready_Hand"
      ProcessValue <- "DIx_DB_Vibro_FB_Ready_Hand"
   Button "Button_44" at 546,92 size 49x22; TextOff 'Выкл'
      on Click: ResetBit("DIx_DB_Vibro_FB_Ready_Start_M")
   Button "Button_45" at 490,92 size 47x22; TextOff 'Вкл'
      on Click: SetBit("DIx_DB_Vibro_FB_Ready_Start_M")
      Appearance <- "DIx_DB_Vibro_FB_Ready_Start_M"
   IOField "I/O field_19" at 666,92 size 23x22; FormatPattern 99
      ProcessValue <- "DIx_DB_Vibro_FB_Ready_Filter_On_SP"
   IOField "I/O field_20" at 689,92 size 23x22; FormatPattern 99
      ProcessValue <- "DIx_DB_Vibro_FB_Ready_Filter_Off_SP"
   Button "Button_46" at 666,69 size 46x20; TextOff 'Inv'
      on Click: InvertBit("DIx_DB_Vibro_FB_Ready_Inverse")
      Appearance <- "DIx_DB_Vibro_FB_Ready_Inverse"
   TextField "Text field_21" at 437,128 size 45x22; Text 'I 1.2'
   TextField "Text field_22" at 482,128 size 112x22; Text 'Пневмотранс.'
   Circle "Circle_21" at 437,151 size 22x22
      Appearance <- "DIx_DB_Transporter_Input"
   Circle "Circle_22" at 460,151 size 22x22
      Appearance <- "DIx_DB_Transporter_Signal"
   Button "Button_47" at 604,129 size 59x44; TextOff 'Авто'; TextList "Hand"
      on Click: InvertBit("DIx_DB_Transporter_Hand")
      Appearance <- "DIx_DB_Transporter_Hand"
      ProcessValue <- "DIx_DB_Transporter_Hand"
   Button "Button_48" at 546,151 size 49x22; TextOff 'Выкл'
      on Click: ResetBit("DIx_DB_Transporter_Start_M")
   Button "Button_49" at 490,151 size 47x22; TextOff 'Вкл'
      on Click: SetBit("DIx_DB_Transporter_Start_M")
      Appearance <- "DIx_DB_Transporter_Start_M"
   IOField "I/O field_21" at 666,151 size 23x22; FormatPattern 99
      ProcessValue <- "DIx_DB_Transporter_Filter_On_SP"
   IOField "I/O field_22" at 689,151 size 23x22; FormatPattern 99
      ProcessValue <- "DIx_DB_Transporter_Filter_Off_SP"
   Button "Button_50" at 666,128 size 46x20; TextOff 'Inv'
      on Click: InvertBit("DIx_DB_Transporter_Inverse")
      Appearance <- "DIx_DB_Transporter_Inverse"
   TextField "Text field_23" at 437,187 size 45x22; Text 'I 1.3'
   TextField "Text field_24" at 482,187 size 128x22; Text 'Жид.доз.Готов.'
   Circle "Circle_23" at 437,210 size 22x22
      Appearance <- "DIx_DB_DL_FB_Ready_Input"
   Circle "Circle_24" at 460,210 size 22x22
      Appearance <- "DIx_DB_DL_FB_Ready_Signal"
   Button "Button_51" at 604,188 size 59x44; TextOff 'Авто'; TextList "Hand"
      on Click: InvertBit("DIx_DB_DL_FB_Ready_Hand")
      Appearance <- "DIx_DB_DL_FB_Ready_Hand"
      ProcessValue <- "DIx_DB_DL_FB_Ready_Hand"
   Button "Button_52" at 546,210 size 49x22; TextOff 'Выкл'
      on Click: ResetBit("DIx_DB_DL_FB_Ready_Start_M")
   Button "Button_53" at 490,210 size 47x22; TextOff 'Вкл'
      on Click: SetBit("DIx_DB_DL_FB_Ready_Start_M")
      Appearance <- "DIx_DB_DL_FB_Ready_Start_M"
   IOField "I/O field_23" at 666,210 size 23x22; FormatPattern 99
      ProcessValue <- "DIx_DB_DL_FB_Ready_Filter_On_SP"
   IOField "I/O field_24" at 689,210 size 23x22; FormatPattern 99
      ProcessValue <- "DIx_DB_DL_FB_Ready_Filter_Off_SP"
   Button "Button_54" at 666,187 size 46x20; TextOff 'Inv'
      on Click: InvertBit("DIx_DB_DL_FB_Ready_Inverse")
      Appearance <- "DIx_DB_DL_FB_Ready_Inverse"
   TextField "Text field_25" at 437,247 size 45x22; Text 'I 1.4'
   TextField "Text field_26" at 482,247 size 61x22; Text 'Проток'
   Circle "Circle_25" at 437,270 size 22x22
      Appearance <- "DIx_DB_Flow_Input"
   Circle "Circle_26" at 460,270 size 22x22
      Appearance <- "DIx_DB_Flow_Signal"
   Button "Button_55" at 604,248 size 59x44; TextOff 'Авто'; TextList "Hand"
      on Click: InvertBit("DIx_DB_Flow_Hand")
      Appearance <- "DIx_DB_Flow_Hand"
      ProcessValue <- "DIx_DB_Flow_Hand"
   Button "Button_56" at 546,270 size 49x22; TextOff 'Выкл'
      on Click: ResetBit("DIx_DB_Flow_Start_M")
   Button "Button_57" at 490,270 size 47x22; TextOff 'Вкл'
      on Click: SetBit("DIx_DB_Flow_Start_M")
      Appearance <- "DIx_DB_Flow_Start_M"
   IOField "I/O field_25" at 666,270 size 23x22; FormatPattern 99
      ProcessValue <- "DIx_DB_Flow_Filter_On_SP"
   IOField "I/O field_26" at 689,270 size 23x22; FormatPattern 99
      ProcessValue <- "DIx_DB_Flow_Filter_Off_SP"
   Button "Button_58" at 666,247 size 46x20; TextOff 'Inv'
      on Click: InvertBit("DIx_DB_Flow_Inverse")
      Appearance <- "DIx_DB_Flow_Inverse"
   TextField "Text field_27" at 437,306 size 45x22; Text 'I 1.5'
   TextField "Text field_28" at 482,306 size 70x22; Text 'Останов'
   Circle "Circle_27" at 437,329 size 22x22
      Appearance <- "DIx_DB_AllBlock_Input"
   Circle "Circle_28" at 460,329 size 22x22
      Appearance <- "DIx_DB_AllBlock_Signal"
   Button "Button_59" at 604,307 size 59x44; TextOff 'Авто'; TextList "Hand"
      on Click: InvertBit("DIx_DB_AllBlock_Hand")
      Appearance <- "DIx_DB_AllBlock_Hand"
      ProcessValue <- "DIx_DB_AllBlock_Hand"
   Button "Button_60" at 546,329 size 49x22; TextOff 'Выкл'
      on Click: ResetBit("DIx_DB_AllBlock_Start_M")
   Button "Button_61" at 490,329 size 47x22; TextOff 'Вкл'
      on Click: SetBit("DIx_DB_AllBlock_Start_M")
      Appearance <- "DIx_DB_AllBlock_Start_M"
   IOField "I/O field_27" at 666,329 size 23x22; FormatPattern 99
      ProcessValue <- "DIx_DB_AllBlock_Filter_On_SP"
   IOField "I/O field_28" at 689,329 size 23x22; FormatPattern 99
      ProcessValue <- "DIx_DB_AllBlock_Filter_Off_SP"
   Button "Button_62" at 666,306 size 46x20; TextOff 'Inv'
      on Click: InvertBit("DIx_DB_AllBlock_Inverse")
      Appearance <- "DIx_DB_AllBlock_Inverse"

screen "DO" 800x480, template "Main"
   Button "Button_1" at 7,5 size 96x32; TextOff 'Мешалки'; Authorization "Admin"
      on Release: ActivateScreen("Mix", 0); SetTag("settings", 1)
      Appearance <- "settings"
   Button "Button_2" at 7,52 size 96x32; TextOff 'Дозаторы'; Authorization "Admin"
      on Release: ActivateScreen("Dos", 0); SetTag("settings", 2)
      Appearance <- "settings"
   Button "Button_3" at 7,99 size 96x32; TextOff 'Клапана'; Authorization "Admin"
      on Release: ActivateScreen("Valve", 0); SetTag("settings", 3)
      Appearance <- "settings"
   Button "Button_4" at 7,146 size 96x32; TextOff 'AI'; Authorization "Admin"
      on Release: ActivateScreen("AI", 0); SetTag("settings", 4)
      Appearance <- "settings"
   Button "Button_5" at 7,193 size 96x32; TextOff 'DI'; Authorization "Admin"
      on Release: ActivateScreen("DI", 0); SetTag("settings", 5)
      Appearance <- "settings"
   Button "Button_6" at 7,240 size 96x32; TextOff 'DO'; Authorization "Admin"
      on Release: ActivateScreen("DO", 0); SetTag("settings", 6)
      Appearance <- "settings"
   Group "Group" at 127,7 size 283x51; TextList "Hand"
   Group "Group_1" at 127,66 size 283x51; TextList "Hand"; Text 'Q 0.0'
   Group "Group_2" at 127,125 size 283x51; TextList "Hand"; Text 'Q 0.0'
   Group "Group_3" at 127,184 size 283x51; TextList "Hand"; Text 'Q 0.0'
   Group "Group_4" at 127,244 size 283x51; TextList "Hand"; Text 'Q 0.0'
   Group "Group_5" at 127,303 size 283x51; TextList "Hand"; Text 'Q 0.0'
   Group "Group_6" at 127,362 size 283x51; TextList "Hand"; Text 'Q 0.0'
   Group "Group_7" at 127,422 size 283x51; TextList "Hand"; Text 'Q 0.0'
   Group "Group_8" at 433,7 size 283x51; TextList "Hand"; Text 'Q 0.0'
   Group "Group_9" at 433,66 size 283x51; Text 'Q 0.0'; TextList "Hand"
   TextField "Text field_4" at 131,10 size 45x22; Text 'Q 0.0'
   TextField "Text field_5" at 176,10 size 69x22; Text 'M1 Пуск'
   Circle "Circle_3" at 131,33 size 22x22
      Appearance <- "DOx_DB_M1_CMD_Start_A"
   Circle "Circle_4" at 154,33 size 22x22
      Appearance <- "DOx_DB_M1_CMD_Q"
   Button "Button_13" at 298,11 size 59x44; TextOff 'Авто'; TextList "Hand"
      on Click: InvertBit("DOx_DB_M1_CMD_Hand")
      Appearance <- "DOx_DB_M1_CMD_Hand"
      ProcessValue <- "DOx_DB_M1_CMD_Hand"
   Button "Button_14" at 240,33 size 49x22; TextOff 'Выкл'
      on Click: ResetBit("DOx_DB_M1_CMD_Start_M")
   Button "Button_15" at 184,33 size 47x22; TextOff 'Вкл'
      on Click: SetBit("DOx_DB_M1_CMD_Start_M")
      Appearance <- "DOx_DB_M1_CMD_Start_M"
   Button "Button_16" at 360,10 size 46x20; TextOff 'Inv'
      on Click: InvertBit("DOx_DB_M1_CMD_Inverse")
      Appearance <- "DOx_DB_M1_CMD_Inverse"
   Button "Button_17" at 360,35 size 46x20; TextOff 'Sim'
      on Click: InvertBit("DOx_DB_M1_CMD_Simulation")
      Appearance <- "DOx_DB_M1_CMD_Simulation"
   TextField "Text field_1" at 131,69 size 45x22; Text 'Q 0.1'
   TextField "Text field_2" at 176,69 size 69x22; Text 'M2 Пуск'
   Circle "Circle_1" at 131,92 size 22x22
      Appearance <- "DOx_DB_M2_CMD_Start_A"
   Circle "Circle_2" at 154,92 size 22x22
      Appearance <- "DOx_DB_M2_CMD_Q"
   Button "Button_7" at 298,70 size 59x44; TextOff 'Авто'; TextList "Hand"
      on Click: InvertBit("DOx_DB_M2_CMD_Hand")
      Appearance <- "DOx_DB_M2_CMD_Hand"
      ProcessValue <- "DOx_DB_M2_CMD_Hand"
   Button "Button_8" at 240,92 size 49x22; TextOff 'Выкл'
      on Click: ResetBit("DOx_DB_M2_CMD_Start_M")
   Button "Button_9" at 184,92 size 47x22; TextOff 'Вкл'
      on Click: SetBit("DOx_DB_M2_CMD_Start_M")
      Appearance <- "DOx_DB_M2_CMD_Start_M"
   Button "Button_10" at 360,69 size 46x20; TextOff 'Inv'
      on Click: InvertBit("DOx_DB_M2_CMD_Inverse")
      Appearance <- "DOx_DB_M2_CMD_Inverse"
   Button "Button_11" at 360,94 size 46x20; TextOff 'Sim'
      on Click: InvertBit("DOx_DB_M2_CMD_Simulation")
      Appearance <- "DOx_DB_M2_CMD_Simulation"
   TextField "Text field_3" at 131,128 size 45x22; Text 'Q 0.2'
   TextField "Text field_6" at 176,128 size 69x22; Text 'M3 Пуск'
   Circle "Circle_5" at 131,151 size 22x22
      Appearance <- "DOx_DB_M3_CMD_Start_A"
   Circle "Circle_6" at 154,151 size 22x22
      Appearance <- "DOx_DB_M3_CMD_Q"
   Button "Button_12" at 298,129 size 59x44; TextOff 'Авто'; TextList "Hand"
      on Click: InvertBit("DOx_DB_M3_CMD_Hand")
      Appearance <- "DOx_DB_M3_CMD_Hand"
      ProcessValue <- "DOx_DB_M3_CMD_Hand"
   Button "Button_18" at 240,151 size 49x22; TextOff 'Выкл'
      on Click: ResetBit("DOx_DB_M3_CMD_Start_M")
   Button "Button_19" at 184,151 size 47x22; TextOff 'Вкл'
      on Click: SetBit("DOx_DB_M3_CMD_Start_M")
      Appearance <- "DOx_DB_M3_CMD_Start_M"
   Button "Button_20" at 360,128 size 46x20; TextOff 'Inv'
      on Click: InvertBit("DOx_DB_M3_CMD_Inverse")
      Appearance <- "DOx_DB_M3_CMD_Inverse"
   Button "Button_21" at 360,153 size 46x20; TextOff 'Sim'
      on Click: InvertBit("DOx_DB_M3_CMD_Simulation")
      Appearance <- "DOx_DB_M3_CMD_Simulation"
   TextField "Text field_7" at 131,187 size 45x22; Text 'Q 0.3'
   TextField "Text field_8" at 176,187 size 109x22; Text 'Сух.Доз.Пуск'
   Circle "Circle_7" at 131,210 size 22x22
      Appearance <- "DOx_DB_DD_CMD_Start_A"
   Circle "Circle_8" at 154,210 size 22x22
      Appearance <- "DOx_DB_DD_CMD_Q"
   Button "Button_22" at 298,188 size 59x44; TextOff 'Авто'; TextList "Hand"
      on Click: InvertBit("DOx_DB_DD_CMD_Hand")
      Appearance <- "DOx_DB_DD_CMD_Hand"
      ProcessValue <- "DOx_DB_DD_CMD_Hand"
   Button "Button_23" at 240,210 size 49x22; TextOff 'Выкл'
      on Click: ResetBit("DOx_DB_DD_CMD_Start_M")
   Button "Button_24" at 184,210 size 47x22; TextOff 'Вкл'
      on Click: SetBit("DOx_DB_DD_CMD_Start_M")